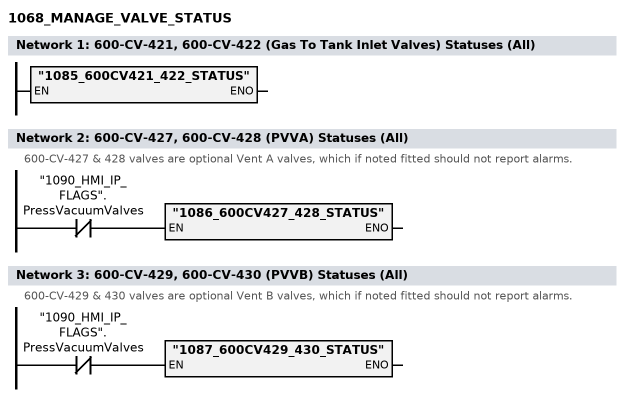
   RUNG wire#powerrail
      "1085_600CV421_422_STATUS"()
   END_RUNG
   // the same network as SCL:
   "1085_600CV421_422_STATUS"();
END_REGION

REGION Network 2: 600-CV-427, 600-CV-428 (PVVA) Statuses (All)
   // 600-CV-427 & 428 valves are optional Vent A valves, which if noted fitted should not report alarms.
   RUNG wire#powerrail
      I_Contact( "1090_HMI_IP_FLAGS".PressVacuumValves )
      "1086_600CV427_428_STATUS"()
   END_RUNG
   // the same network as SCL:
   IF NOT "1090_HMI_IP_FLAGS".PressVacuumValves THEN "1086_600CV427_428_STATUS"(); END_IF;
END_REGION

REGION Network 3: 600-CV-429, 600-CV-430 (PVVB) Statuses (All)
   // 600-CV-429 & 430 valves are optional Vent B valves, which if noted fitted should not report alarms.
   RUNG wire#powerrail
      I_Contact( "1090_HMI_IP_FLAGS".PressVacuumValves )
      "1087_600CV429_430_STATUS"()
   END_RUNG
   // the same network as SCL:
   IF NOT "1090_HMI_IP_FLAGS".PressVacuumValves THEN "1087_600CV429_430_STATUS"(); END_IF;
END_REGION
END_FUNCTION

// folder: 1000 - 1999 BWT System Control/1060 - 1089 Alarm & Valve Status Handling/1070 - 1079 Tank Alarms

FUNCTION "1070_LT421_422_ALARMS" : Void   // FC1070, LAD
{ S7_Optimized_Access := 'TRUE' }
VERSION : 0.1
// Alarm wrapper function for BWT Level on each tank.
// DummyIn and DummyAlarm are used to manage the unused I/O in the analog health trips function as this function only uses Low and High warnings, it does not output HighHigh or LowLow alarms.
   VAR_TEMP
      DummyIn : Real;   // Dummy input used if alarms are Low and High only.
      DummyAlarm : Bool;   // Dummy output used if alarms are Low and High only.
   END_VAR
BEGIN

REGION Network 1: LT421, LT422 Alarms (RIO 01: FPT. 1P, 1S)
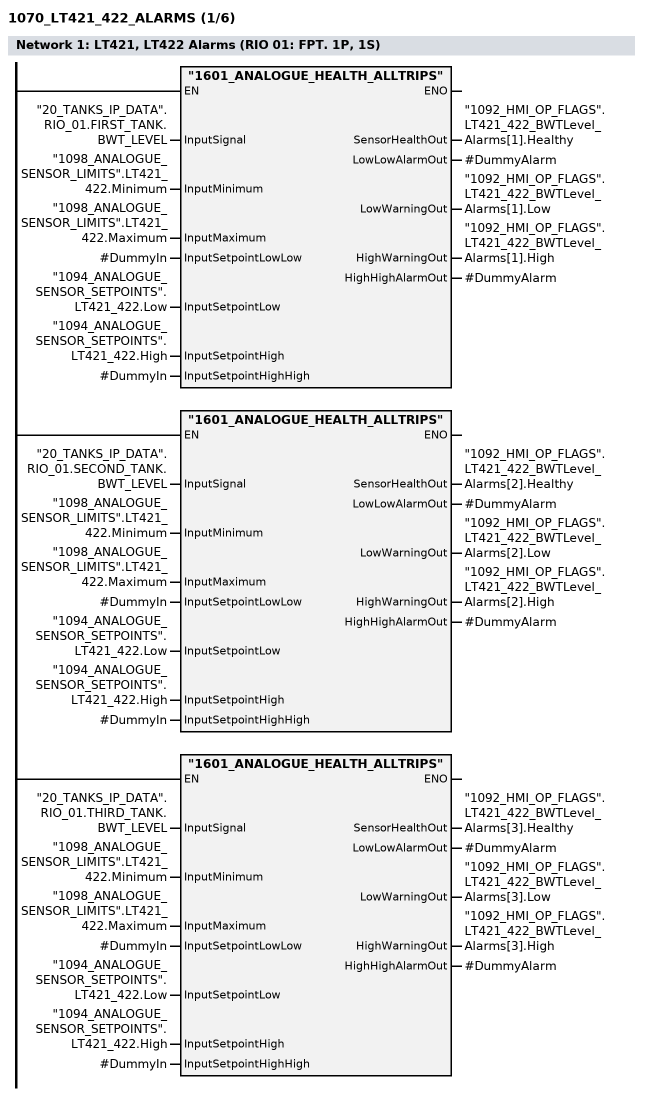
   RUNG wire#powerrail
      "1601_ANALOGUE_HEALTH_ALLTRIPS"(InputSignal := "20_TANKS_IP_DATA".RIO_01.FIRST_TANK.BWT_LEVEL, InputMinimum := "1098_ANALOGUE_SENSOR_LIMITS".LT421_422.Minimum, InputMaximum := "1098_ANALOGUE_SENSOR_LIMITS".LT421_422.Maximum, InputSetpointLowLow := #DummyIn, InputSetpointLow := "1094_ANALOGUE_SENSOR_SETPOINTS".LT421_422.Low, InputSetpointHigh := "1094_ANALOGUE_SENSOR_SETPOINTS".LT421_422.High, InputSetpointHighHigh := #DummyIn, SensorHealthOut => "1092_HMI_OP_FLAGS".LT421_422_BWTLevel_Alarms[1].Healthy, LowLowAlarmOut => #DummyAlarm, LowWarningOut => "1092_HMI_OP_FLAGS".LT421_422_BWTLevel_Alarms[1].Low, HighWarningOut => "1092_HMI_OP_FLAGS".LT421_422_BWTLevel_Alarms[1].High, HighHighAlarmOut => #DummyAlarm)
   END_RUNG
   RUNG wire#powerrail
      "1601_ANALOGUE_HEALTH_ALLTRIPS"(InputSignal := "20_TANKS_IP_DATA".RIO_01.SECOND_TANK.BWT_LEVEL, InputMinimum := "1098_ANALOGUE_SENSOR_LIMITS".LT421_422.Minimum, InputMaximum := "1098_ANALOGUE_SENSOR_LIMITS".LT421_422.Maximum, InputSetpointLowLow := #DummyIn, InputSetpointLow := "1094_ANALOGUE_SENSOR_SETPOINTS".LT421_422.Low, InputSetpointHigh := "1094_ANALOGUE_SENSOR_SETPOINTS".LT421_422.High, InputSetpointHighHigh := #DummyIn, SensorHealthOut => "1092_HMI_OP_FLAGS".LT421_422_BWTLevel_Alarms[2].Healthy, LowLowAlarmOut => #DummyAlarm, LowWarningOut => "1092_HMI_OP_FLAGS".LT421_422_BWTLevel_Alarms[2].Low, HighWarningOut => "1092_HMI_OP_FLAGS".LT421_422_BWTLevel_Alarms[2].High, HighHighAlarmOut => #DummyAlarm)
   END_RUNG
   RUNG wire#powerrail
      "1601_ANALOGUE_HEALTH_ALLTRIPS"(InputSignal := "20_TANKS_IP_DATA".RIO_01.THIRD_TANK.BWT_LEVEL, InputMinimum := "1098_ANALOGUE_SENSOR_LIMITS".LT421_422.Minimum, InputMaximum := "1098_ANALOGUE_SENSOR_LIMITS".LT421_422.Maximum, InputSetpointLowLow := #DummyIn, InputSetpointLow := "1094_ANALOGUE_SENSOR_SETPOINTS".LT421_422.Low, InputSetpointHigh := "1094_ANALOGUE_SENSOR_SETPOINTS".LT421_422.High, InputSetpointHighHigh := #DummyIn, SensorHealthOut => "1092_HMI_OP_FLAGS".LT421_422_BWTLevel_Alarms[3].Healthy, LowLowAlarmOut => #DummyAlarm, LowWarningOut => "1092_HMI_OP_FLAGS".LT421_422_BWTLevel_Alarms[3].Low, HighWarningOut => "1092_HMI_OP_FLAGS".LT421_422_BWTLevel_Alarms[3].High, HighHighAlarmOut => #DummyAlarm)
   END_RUNG
   // the same network as SCL:
   "1601_ANALOGUE_HEALTH_ALLTRIPS"(InputSignal := "20_TANKS_IP_DATA".RIO_01.FIRST_TANK.BWT_LEVEL,
                           InputMinimum := "1098_ANALOGUE_SENSOR_LIMITS".LT421_422.Minimum,
                           InputMaximum := "1098_ANALOGUE_SENSOR_LIMITS".LT421_422.Maximum,
                           InputSetpointLowLow := #DummyIn,
                           InputSetpointLow := "1094_ANALOGUE_SENSOR_SETPOINTS".LT421_422.Low,
                           InputSetpointHigh := "1094_ANALOGUE_SENSOR_SETPOINTS".LT421_422.High,
                           InputSetpointHighHigh := #DummyIn,
                           SensorHealthOut => "1092_HMI_OP_FLAGS".LT421_422_BWTLevel_Alarms[1].Healthy,
                           LowLowAlarmOut => #DummyAlarm,
                           LowWarningOut => "1092_HMI_OP_FLAGS".LT421_422_BWTLevel_Alarms[1].Low,
                           HighWarningOut => "1092_HMI_OP_FLAGS".LT421_422_BWTLevel_Alarms[1].High,
                           HighHighAlarmOut => #DummyAlarm);
   "1601_ANALOGUE_HEALTH_ALLTRIPS"(InputSignal := "20_TANKS_IP_DATA".RIO_01.SECOND_TANK.BWT_LEVEL,
                           InputMinimum := "1098_ANALOGUE_SENSOR_LIMITS".LT421_422.Minimum,
                           InputMaximum := "1098_ANALOGUE_SENSOR_LIMITS".LT421_422.Maximum,
                           InputSetpointLowLow := #DummyIn,
                           InputSetpointLow := "1094_ANALOGUE_SENSOR_SETPOINTS".LT421_422.Low,
                           InputSetpointHigh := "1094_ANALOGUE_SENSOR_SETPOINTS".LT421_422.High,
                           InputSetpointHighHigh := #DummyIn,
                           SensorHealthOut => "1092_HMI_OP_FLAGS".LT421_422_BWTLevel_Alarms[2].Healthy,
                           LowLowAlarmOut => #DummyAlarm,
                           LowWarningOut => "1092_HMI_OP_FLAGS".LT421_422_BWTLevel_Alarms[2].Low,
                           HighWarningOut => "1092_HMI_OP_FLAGS".LT421_422_BWTLevel_Alarms[2].High,
                           HighHighAlarmOut => #DummyAlarm);
   "1601_ANALOGUE_HEALTH_ALLTRIPS"(InputSignal := "20_TANKS_IP_DATA".RIO_01.THIRD_TANK.BWT_LEVEL,
                           InputMinimum := "1098_ANALOGUE_SENSOR_LIMITS".LT421_422.Minimum,
                           InputMaximum := "1098_ANALOGUE_SENSOR_LIMITS".LT421_422.Maximum,
                           InputSetpointLowLow := #DummyIn,
                           InputSetpointLow := "1094_ANALOGUE_SENSOR_SETPOINTS".LT421_422.Low,
                           InputSetpointHigh := "1094_ANALOGUE_SENSOR_SETPOINTS".LT421_422.High,
                           InputSetpointHighHigh := #DummyIn,
                           SensorHealthOut => "1092_HMI_OP_FLAGS".LT421_422_BWTLevel_Alarms[3].Healthy,
                           LowLowAlarmOut => #DummyAlarm,
                           LowWarningOut => "1092_HMI_OP_FLAGS".LT421_422_BWTLevel_Alarms[3].Low,
                           HighWarningOut => "1092_HMI_OP_FLAGS".LT421_422_BWTLevel_Alarms[3].High,
                           HighHighAlarmOut => #DummyAlarm);
END_REGION

REGION Network 2: LT421, LT422 Alarms (RIO 02: 2P, 2S)
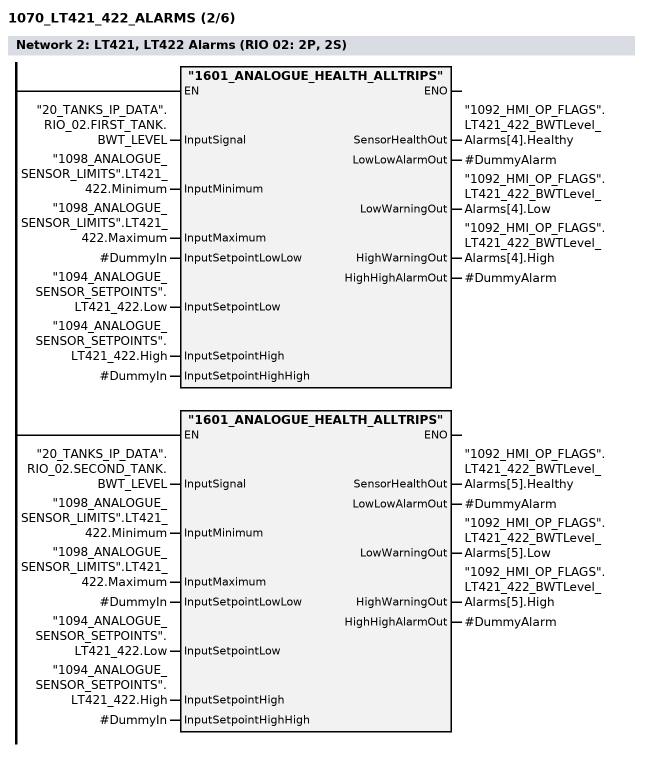
   RUNG wire#powerrail
      "1601_ANALOGUE_HEALTH_ALLTRIPS"(InputSignal := "20_TANKS_IP_DATA".RIO_02.FIRST_TANK.BWT_LEVEL, InputMinimum := "1098_ANALOGUE_SENSOR_LIMITS".LT421_422.Minimum, InputMaximum := "1098_ANALOGUE_SENSOR_LIMITS".LT421_422.Maximum, InputSetpointLowLow := #DummyIn, InputSetpointLow := "1094_ANALOGUE_SENSOR_SETPOINTS".LT421_422.Low, InputSetpointHigh := "1094_ANALOGUE_SENSOR_SETPOINTS".LT421_422.High, InputSetpointHighHigh := #DummyIn, SensorHealthOut => "1092_HMI_OP_FLAGS".LT421_422_BWTLevel_Alarms[4].Healthy, LowLowAlarmOut => #DummyAlarm, LowWarningOut => "1092_HMI_OP_FLAGS".LT421_422_BWTLevel_Alarms[4].Low, HighWarningOut => "1092_HMI_OP_FLAGS".LT421_422_BWTLevel_Alarms[4].High, HighHighAlarmOut => #DummyAlarm)
   END_RUNG
   RUNG wire#powerrail
      "1601_ANALOGUE_HEALTH_ALLTRIPS"(InputSignal := "20_TANKS_IP_DATA".RIO_02.SECOND_TANK.BWT_LEVEL, InputMinimum := "1098_ANALOGUE_SENSOR_LIMITS".LT421_422.Minimum, InputMaximum := "1098_ANALOGUE_SENSOR_LIMITS".LT421_422.Maximum, InputSetpointLowLow := #DummyIn, InputSetpointLow := "1094_ANALOGUE_SENSOR_SETPOINTS".LT421_422.Low, InputSetpointHigh := "1094_ANALOGUE_SENSOR_SETPOINTS".LT421_422.High, InputSetpointHighHigh := #DummyIn, SensorHealthOut => "1092_HMI_OP_FLAGS".LT421_422_BWTLevel_Alarms[5].Healthy, LowLowAlarmOut => #DummyAlarm, LowWarningOut => "1092_HMI_OP_FLAGS".LT421_422_BWTLevel_Alarms[5].Low, HighWarningOut => "1092_HMI_OP_FLAGS".LT421_422_BWTLevel_Alarms[5].High, HighHighAlarmOut => #DummyAlarm)
   END_RUNG
   // the same network as SCL:
   "1601_ANALOGUE_HEALTH_ALLTRIPS"(InputSignal := "20_TANKS_IP_DATA".RIO_02.FIRST_TANK.BWT_LEVEL,
                           InputMinimum := "1098_ANALOGUE_SENSOR_LIMITS".LT421_422.Minimum,
                           InputMaximum := "1098_ANALOGUE_SENSOR_LIMITS".LT421_422.Maximum,
                           InputSetpointLowLow := #DummyIn,
                           InputSetpointLow := "1094_ANALOGUE_SENSOR_SETPOINTS".LT421_422.Low,
                           InputSetpointHigh := "1094_ANALOGUE_SENSOR_SETPOINTS".LT421_422.High,
                           InputSetpointHighHigh := #DummyIn,
                           SensorHealthOut => "1092_HMI_OP_FLAGS".LT421_422_BWTLevel_Alarms[4].Healthy,
                           LowLowAlarmOut => #DummyAlarm,
                           LowWarningOut => "1092_HMI_OP_FLAGS".LT421_422_BWTLevel_Alarms[4].Low,
                           HighWarningOut => "1092_HMI_OP_FLAGS".LT421_422_BWTLevel_Alarms[4].High,
                           HighHighAlarmOut => #DummyAlarm);
   "1601_ANALOGUE_HEALTH_ALLTRIPS"(InputSignal := "20_TANKS_IP_DATA".RIO_02.SECOND_TANK.BWT_LEVEL,
                           InputMinimum := "1098_ANALOGUE_SENSOR_LIMITS".LT421_422.Minimum,
                           InputMaximum := "1098_ANALOGUE_SENSOR_LIMITS".LT421_422.Maximum,
                           InputSetpointLowLow := #DummyIn,
                           InputSetpointLow := "1094_ANALOGUE_SENSOR_SETPOINTS".LT421_422.Low,
                           InputSetpointHigh := "1094_ANALOGUE_SENSOR_SETPOINTS".LT421_422.High,
                           InputSetpointHighHigh := #DummyIn,
                           SensorHealthOut => "1092_HMI_OP_FLAGS".LT421_422_BWTLevel_Alarms[5].Healthy,
                           LowLowAlarmOut => #DummyAlarm,
                           LowWarningOut => "1092_HMI_OP_FLAGS".LT421_422_BWTLevel_Alarms[5].Low,
                           HighWarningOut => "1092_HMI_OP_FLAGS".LT421_422_BWTLevel_Alarms[5].High,
                           HighHighAlarmOut => #DummyAlarm);
END_REGION

REGION Network 3: LT421, LT422 Alarms (RIO 03: 3P, 3S)
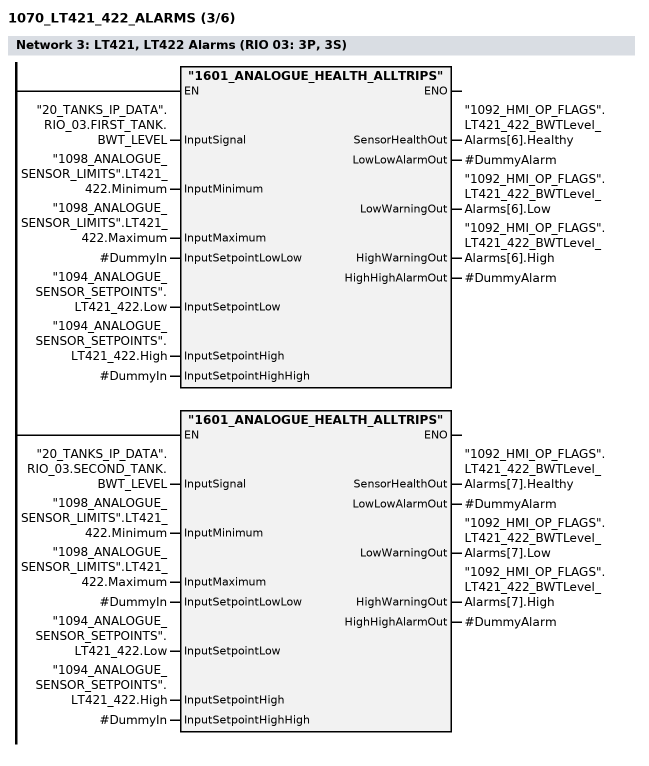
   RUNG wire#powerrail
      "1601_ANALOGUE_HEALTH_ALLTRIPS"(InputSignal := "20_TANKS_IP_DATA".RIO_03.FIRST_TANK.BWT_LEVEL, InputMinimum := "1098_ANALOGUE_SENSOR_LIMITS".LT421_422.Minimum, InputMaximum := "1098_ANALOGUE_SENSOR_LIMITS".LT421_422.Maximum, InputSetpointLowLow := #DummyIn, InputSetpointLow := "1094_ANALOGUE_SENSOR_SETPOINTS".LT421_422.Low, InputSetpointHigh := "1094_ANALOGUE_SENSOR_SETPOINTS".LT421_422.High, InputSetpointHighHigh := #DummyIn, SensorHealthOut => "1092_HMI_OP_FLAGS".LT421_422_BWTLevel_Alarms[6].Healthy, LowLowAlarmOut => #DummyAlarm, LowWarningOut => "1092_HMI_OP_FLAGS".LT421_422_BWTLevel_Alarms[6].Low, HighWarningOut => "1092_HMI_OP_FLAGS".LT421_422_BWTLevel_Alarms[6].High, HighHighAlarmOut => #DummyAlarm)
   END_RUNG
   RUNG wire#powerrail
      "1601_ANALOGUE_HEALTH_ALLTRIPS"(InputSignal := "20_TANKS_IP_DATA".RIO_03.SECOND_TANK.BWT_LEVEL, InputMinimum := "1098_ANALOGUE_SENSOR_LIMITS".LT421_422.Minimum, InputMaximum := "1098_ANALOGUE_SENSOR_LIMITS".LT421_422.Maximum, InputSetpointLowLow := #DummyIn, InputSetpointLow := "1094_ANALOGUE_SENSOR_SETPOINTS".LT421_422.Low, InputSetpointHigh := "1094_ANALOGUE_SENSOR_SETPOINTS".LT421_422.High, InputSetpointHighHigh := #DummyIn, SensorHealthOut => "1092_HMI_OP_FLAGS".LT421_422_BWTLevel_Alarms[7].Healthy, LowLowAlarmOut => #DummyAlarm, LowWarningOut => "1092_HMI_OP_FLAGS".LT421_422_BWTLevel_Alarms[7].Low, HighWarningOut => "1092_HMI_OP_FLAGS".LT421_422_BWTLevel_Alarms[7].High, HighHighAlarmOut => #DummyAlarm)
   END_RUNG
   // the same network as SCL:
   "1601_ANALOGUE_HEALTH_ALLTRIPS"(InputSignal := "20_TANKS_IP_DATA".RIO_03.FIRST_TANK.BWT_LEVEL,
                           InputMinimum := "1098_ANALOGUE_SENSOR_LIMITS".LT421_422.Minimum,
                           InputMaximum := "1098_ANALOGUE_SENSOR_LIMITS".LT421_422.Maximum,
                           InputSetpointLowLow := #DummyIn,
                           InputSetpointLow := "1094_ANALOGUE_SENSOR_SETPOINTS".LT421_422.Low,
                           InputSetpointHigh := "1094_ANALOGUE_SENSOR_SETPOINTS".LT421_422.High,
                           InputSetpointHighHigh := #DummyIn,
                           SensorHealthOut => "1092_HMI_OP_FLAGS".LT421_422_BWTLevel_Alarms[6].Healthy,
                           LowLowAlarmOut => #DummyAlarm,
                           LowWarningOut => "1092_HMI_OP_FLAGS".LT421_422_BWTLevel_Alarms[6].Low,
                           HighWarningOut => "1092_HMI_OP_FLAGS".LT421_422_BWTLevel_Alarms[6].High,
                           HighHighAlarmOut => #DummyAlarm);
   "1601_ANALOGUE_HEALTH_ALLTRIPS"(InputSignal := "20_TANKS_IP_DATA".RIO_03.SECOND_TANK.BWT_LEVEL,
                           InputMinimum := "1098_ANALOGUE_SENSOR_LIMITS".LT421_422.Minimum,
                           InputMaximum := "1098_ANALOGUE_SENSOR_LIMITS".LT421_422.Maximum,
                           InputSetpointLowLow := #DummyIn,
                           InputSetpointLow := "1094_ANALOGUE_SENSOR_SETPOINTS".LT421_422.Low,
                           InputSetpointHigh := "1094_ANALOGUE_SENSOR_SETPOINTS".LT421_422.High,
                           InputSetpointHighHigh := #DummyIn,
                           SensorHealthOut => "1092_HMI_OP_FLAGS".LT421_422_BWTLevel_Alarms[7].Healthy,
                           LowLowAlarmOut => #DummyAlarm,
                           LowWarningOut => "1092_HMI_OP_FLAGS".LT421_422_BWTLevel_Alarms[7].Low,
                           HighWarningOut => "1092_HMI_OP_FLAGS".LT421_422_BWTLevel_Alarms[7].High,
                           HighHighAlarmOut => #DummyAlarm);
END_REGION

REGION Network 4: LT421, LT422 Alarms (RIO 04: 4P, 4S)
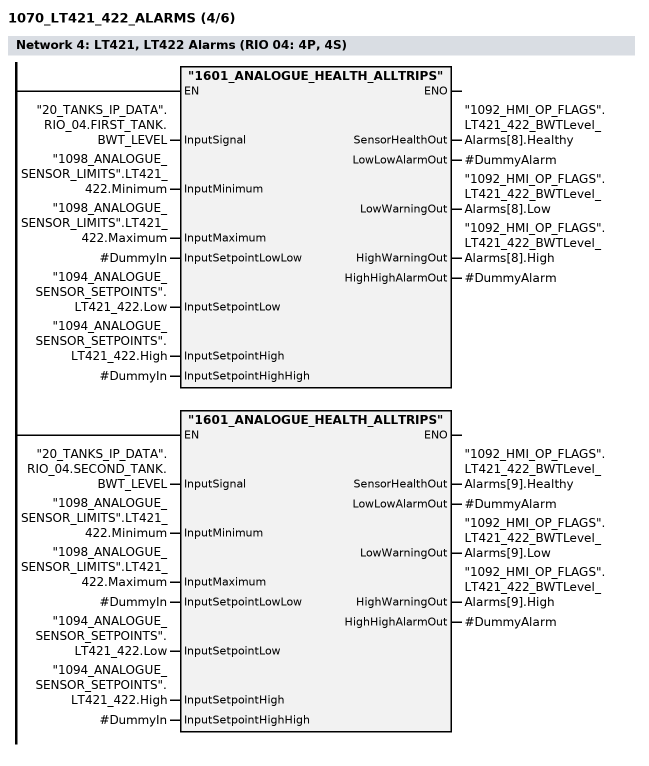
   RUNG wire#powerrail
      "1601_ANALOGUE_HEALTH_ALLTRIPS"(InputSignal := "20_TANKS_IP_DATA".RIO_04.FIRST_TANK.BWT_LEVEL, InputMinimum := "1098_ANALOGUE_SENSOR_LIMITS".LT421_422.Minimum, InputMaximum := "1098_ANALOGUE_SENSOR_LIMITS".LT421_422.Maximum, InputSetpointLowLow := #DummyIn, InputSetpointLow := "1094_ANALOGUE_SENSOR_SETPOINTS".LT421_422.Low, InputSetpointHigh := "1094_ANALOGUE_SENSOR_SETPOINTS".LT421_422.High, InputSetpointHighHigh := #DummyIn, SensorHealthOut => "1092_HMI_OP_FLAGS".LT421_422_BWTLevel_Alarms[8].Healthy, LowLowAlarmOut => #DummyAlarm, LowWarningOut => "1092_HMI_OP_FLAGS".LT421_422_BWTLevel_Alarms[8].Low, HighWarningOut => "1092_HMI_OP_FLAGS".LT421_422_BWTLevel_Alarms[8].High, HighHighAlarmOut => #DummyAlarm)
   END_RUNG
   RUNG wire#powerrail
      "1601_ANALOGUE_HEALTH_ALLTRIPS"(InputSignal := "20_TANKS_IP_DATA".RIO_04.SECOND_TANK.BWT_LEVEL, InputMinimum := "1098_ANALOGUE_SENSOR_LIMITS".LT421_422.Minimum, InputMaximum := "1098_ANALOGUE_SENSOR_LIMITS".LT421_422.Maximum, InputSetpointLowLow := #DummyIn, InputSetpointLow := "1094_ANALOGUE_SENSOR_SETPOINTS".LT421_422.Low, InputSetpointHigh := "1094_ANALOGUE_SENSOR_SETPOINTS".LT421_422.High, InputSetpointHighHigh := #DummyIn, SensorHealthOut => "1092_HMI_OP_FLAGS".LT421_422_BWTLevel_Alarms[9].Healthy, LowLowAlarmOut => #DummyAlarm, LowWarningOut => "1092_HMI_OP_FLAGS".LT421_422_BWTLevel_Alarms[9].Low, HighWarningOut => "1092_HMI_OP_FLAGS".LT421_422_BWTLevel_Alarms[9].High, HighHighAlarmOut => #DummyAlarm)
   END_RUNG
   // the same network as SCL:
   "1601_ANALOGUE_HEALTH_ALLTRIPS"(InputSignal := "20_TANKS_IP_DATA".RIO_04.FIRST_TANK.BWT_LEVEL,
                           InputMinimum := "1098_ANALOGUE_SENSOR_LIMITS".LT421_422.Minimum,
                           InputMaximum := "1098_ANALOGUE_SENSOR_LIMITS".LT421_422.Maximum,
                           InputSetpointLowLow := #DummyIn,
                           InputSetpointLow := "1094_ANALOGUE_SENSOR_SETPOINTS".LT421_422.Low,
                           InputSetpointHigh := "1094_ANALOGUE_SENSOR_SETPOINTS".LT421_422.High,
                           InputSetpointHighHigh := #DummyIn,
                           SensorHealthOut => "1092_HMI_OP_FLAGS".LT421_422_BWTLevel_Alarms[8].Healthy,
                           LowLowAlarmOut => #DummyAlarm,
                           LowWarningOut => "1092_HMI_OP_FLAGS".LT421_422_BWTLevel_Alarms[8].Low,
                           HighWarningOut => "1092_HMI_OP_FLAGS".LT421_422_BWTLevel_Alarms[8].High,
                           HighHighAlarmOut => #DummyAlarm);
   "1601_ANALOGUE_HEALTH_ALLTRIPS"(InputSignal := "20_TANKS_IP_DATA".RIO_04.SECOND_TANK.BWT_LEVEL,
                           InputMinimum := "1098_ANALOGUE_SENSOR_LIMITS".LT421_422.Minimum,
                           InputMaximum := "1098_ANALOGUE_SENSOR_LIMITS".LT421_422.Maximum,
                           InputSetpointLowLow := #DummyIn,
                           InputSetpointLow := "1094_ANALOGUE_SENSOR_SETPOINTS".LT421_422.Low,
                           InputSetpointHigh := "1094_ANALOGUE_SENSOR_SETPOINTS".LT421_422.High,
                           InputSetpointHighHigh := #DummyIn,
                           SensorHealthOut => "1092_HMI_OP_FLAGS".LT421_422_BWTLevel_Alarms[9].Healthy,
                           LowLowAlarmOut => #DummyAlarm,
                           LowWarningOut => "1092_HMI_OP_FLAGS".LT421_422_BWTLevel_Alarms[9].Low,
                           HighWarningOut => "1092_HMI_OP_FLAGS".LT421_422_BWTLevel_Alarms[9].High,
                           HighHighAlarmOut => #DummyAlarm);
END_REGION

REGION Network 5: LT421, LT422 Alarms (RIO 05: 5P, 5S)
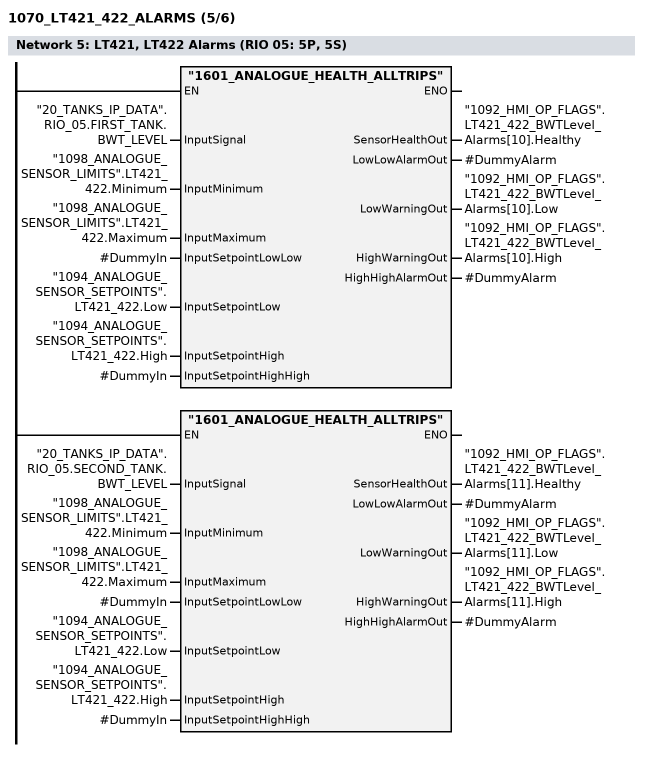
   RUNG wire#powerrail
      "1601_ANALOGUE_HEALTH_ALLTRIPS"(InputSignal := "20_TANKS_IP_DATA".RIO_05.FIRST_TANK.BWT_LEVEL, InputMinimum := "1098_ANALOGUE_SENSOR_LIMITS".LT421_422.Minimum, InputMaximum := "1098_ANALOGUE_SENSOR_LIMITS".LT421_422.Maximum, InputSetpointLowLow := #DummyIn, InputSetpointLow := "1094_ANALOGUE_SENSOR_SETPOINTS".LT421_422.Low, InputSetpointHigh := "1094_ANALOGUE_SENSOR_SETPOINTS".LT421_422.High, InputSetpointHighHigh := #DummyIn, SensorHealthOut => "1092_HMI_OP_FLAGS".LT421_422_BWTLevel_Alarms[10].Healthy, LowLowAlarmOut => #DummyAlarm, LowWarningOut => "1092_HMI_OP_FLAGS".LT421_422_BWTLevel_Alarms[10].Low, HighWarningOut => "1092_HMI_OP_FLAGS".LT421_422_BWTLevel_Alarms[10].High, HighHighAlarmOut => #DummyAlarm)
   END_RUNG
   RUNG wire#powerrail
      "1601_ANALOGUE_HEALTH_ALLTRIPS"(InputSignal := "20_TANKS_IP_DATA".RIO_05.SECOND_TANK.BWT_LEVEL, InputMinimum := "1098_ANALOGUE_SENSOR_LIMITS".LT421_422.Minimum, InputMaximum := "1098_ANALOGUE_SENSOR_LIMITS".LT421_422.Maximum, InputSetpointLowLow := #DummyIn, InputSetpointLow := "1094_ANALOGUE_SENSOR_SETPOINTS".LT421_422.Low, InputSetpointHigh := "1094_ANALOGUE_SENSOR_SETPOINTS".LT421_422.High, InputSetpointHighHigh := #DummyIn, SensorHealthOut => "1092_HMI_OP_FLAGS".LT421_422_BWTLevel_Alarms[11].Healthy, LowLowAlarmOut => #DummyAlarm, LowWarningOut => "1092_HMI_OP_FLAGS".LT421_422_BWTLevel_Alarms[11].Low, HighWarningOut => "1092_HMI_OP_FLAGS".LT421_422_BWTLevel_Alarms[11].High, HighHighAlarmOut => #DummyAlarm)
   END_RUNG
   // the same network as SCL:
   "1601_ANALOGUE_HEALTH_ALLTRIPS"(InputSignal := "20_TANKS_IP_DATA".RIO_05.FIRST_TANK.BWT_LEVEL,
                           InputMinimum := "1098_ANALOGUE_SENSOR_LIMITS".LT421_422.Minimum,
                           InputMaximum := "1098_ANALOGUE_SENSOR_LIMITS".LT421_422.Maximum,
                           InputSetpointLowLow := #DummyIn,
                           InputSetpointLow := "1094_ANALOGUE_SENSOR_SETPOINTS".LT421_422.Low,
                           InputSetpointHigh := "1094_ANALOGUE_SENSOR_SETPOINTS".LT421_422.High,
                           InputSetpointHighHigh := #DummyIn,
                           SensorHealthOut => "1092_HMI_OP_FLAGS".LT421_422_BWTLevel_Alarms[10].Healthy,
                           LowLowAlarmOut => #DummyAlarm,
                           LowWarningOut => "1092_HMI_OP_FLAGS".LT421_422_BWTLevel_Alarms[10].Low,
                           HighWarningOut => "1092_HMI_OP_FLAGS".LT421_422_BWTLevel_Alarms[10].High,
                           HighHighAlarmOut => #DummyAlarm);
   "1601_ANALOGUE_HEALTH_ALLTRIPS"(InputSignal := "20_TANKS_IP_DATA".RIO_05.SECOND_TANK.BWT_LEVEL,
                           InputMinimum := "1098_ANALOGUE_SENSOR_LIMITS".LT421_422.Minimum,
                           InputMaximum := "1098_ANALOGUE_SENSOR_LIMITS".LT421_422.Maximum,
                           InputSetpointLowLow := #DummyIn,
                           InputSetpointLow := "1094_ANALOGUE_SENSOR_SETPOINTS".LT421_422.Low,
                           InputSetpointHigh := "1094_ANALOGUE_SENSOR_SETPOINTS".LT421_422.High,
                           InputSetpointHighHigh := #DummyIn,
                           SensorHealthOut => "1092_HMI_OP_FLAGS".LT421_422_BWTLevel_Alarms[11].Healthy,
                           LowLowAlarmOut => #DummyAlarm,
                           LowWarningOut => "1092_HMI_OP_FLAGS".LT421_422_BWTLevel_Alarms[11].Low,
                           HighWarningOut => "1092_HMI_OP_FLAGS".LT421_422_BWTLevel_Alarms[11].High,
                           HighHighAlarmOut => #DummyAlarm);
END_REGION

REGION Network 6: LT421, LT422 Alarms (RIO 06: 6P, 6S)
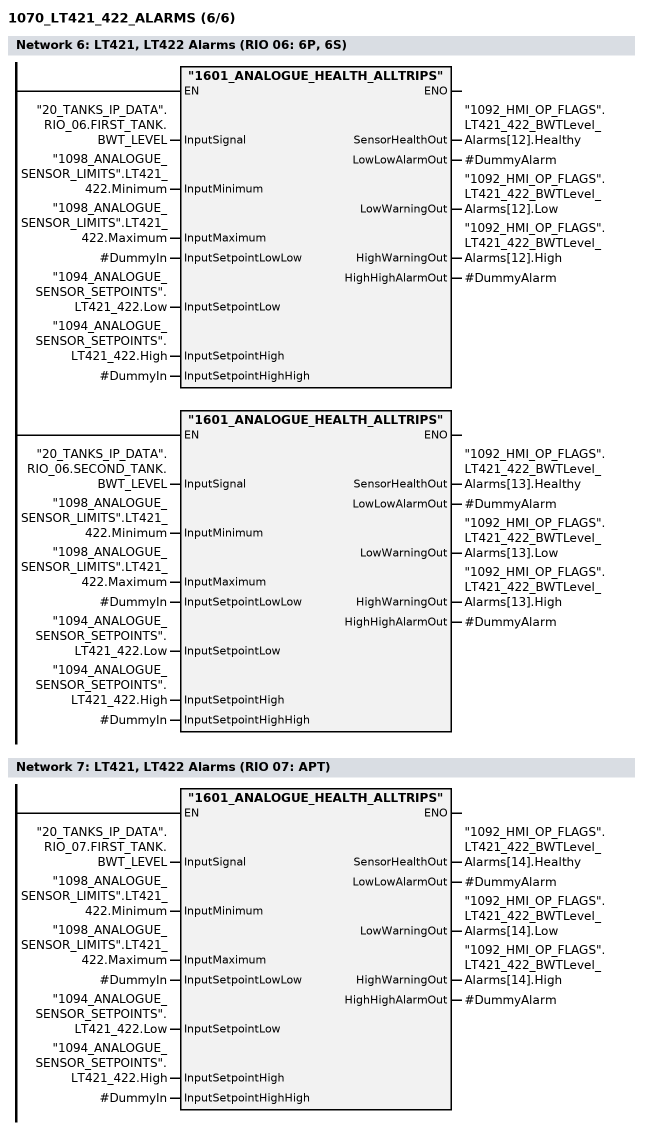
   RUNG wire#powerrail
      "1601_ANALOGUE_HEALTH_ALLTRIPS"(InputSignal := "20_TANKS_IP_DATA".RIO_06.FIRST_TANK.BWT_LEVEL, InputMinimum := "1098_ANALOGUE_SENSOR_LIMITS".LT421_422.Minimum, InputMaximum := "1098_ANALOGUE_SENSOR_LIMITS".LT421_422.Maximum, InputSetpointLowLow := #DummyIn, InputSetpointLow := "1094_ANALOGUE_SENSOR_SETPOINTS".LT421_422.Low, InputSetpointHigh := "1094_ANALOGUE_SENSOR_SETPOINTS".LT421_422.High, InputSetpointHighHigh := #DummyIn, SensorHealthOut => "1092_HMI_OP_FLAGS".LT421_422_BWTLevel_Alarms[12].Healthy, LowLowAlarmOut => #DummyAlarm, LowWarningOut => "1092_HMI_OP_FLAGS".LT421_422_BWTLevel_Alarms[12].Low, HighWarningOut => "1092_HMI_OP_FLAGS".LT421_422_BWTLevel_Alarms[12].High, HighHighAlarmOut => #DummyAlarm)
   END_RUNG
   RUNG wire#powerrail
      "1601_ANALOGUE_HEALTH_ALLTRIPS"(InputSignal := "20_TANKS_IP_DATA".RIO_06.SECOND_TANK.BWT_LEVEL, InputMinimum := "1098_ANALOGUE_SENSOR_LIMITS".LT421_422.Minimum, InputMaximum := "1098_ANALOGUE_SENSOR_LIMITS".LT421_422.Maximum, InputSetpointLowLow := #DummyIn, InputSetpointLow := "1094_ANALOGUE_SENSOR_SETPOINTS".LT421_422.Low, InputSetpointHigh := "1094_ANALOGUE_SENSOR_SETPOINTS".LT421_422.High, InputSetpointHighHigh := #DummyIn, SensorHealthOut => "1092_HMI_OP_FLAGS".LT421_422_BWTLevel_Alarms[13].Healthy, LowLowAlarmOut => #DummyAlarm, LowWarningOut => "1092_HMI_OP_FLAGS".LT421_422_BWTLevel_Alarms[13].Low, HighWarningOut => "1092_HMI_OP_FLAGS".LT421_422_BWTLevel_Alarms[13].High, HighHighAlarmOut => #DummyAlarm)
   END_RUNG
   // the same network as SCL:
   "1601_ANALOGUE_HEALTH_ALLTRIPS"(InputSignal := "20_TANKS_IP_DATA".RIO_06.FIRST_TANK.BWT_LEVEL,
                           InputMinimum := "1098_ANALOGUE_SENSOR_LIMITS".LT421_422.Minimum,
                           InputMaximum := "1098_ANALOGUE_SENSOR_LIMITS".LT421_422.Maximum,
                           InputSetpointLowLow := #DummyIn,
                           InputSetpointLow := "1094_ANALOGUE_SENSOR_SETPOINTS".LT421_422.Low,
                           InputSetpointHigh := "1094_ANALOGUE_SENSOR_SETPOINTS".LT421_422.High,
                           InputSetpointHighHigh := #DummyIn,
                           SensorHealthOut => "1092_HMI_OP_FLAGS".LT421_422_BWTLevel_Alarms[12].Healthy,
                           LowLowAlarmOut => #DummyAlarm,
                           LowWarningOut => "1092_HMI_OP_FLAGS".LT421_422_BWTLevel_Alarms[12].Low,
                           HighWarningOut => "1092_HMI_OP_FLAGS".LT421_422_BWTLevel_Alarms[12].High,
                           HighHighAlarmOut => #DummyAlarm);
   "1601_ANALOGUE_HEALTH_ALLTRIPS"(InputSignal := "20_TANKS_IP_DATA".RIO_06.SECOND_TANK.BWT_LEVEL,
                           InputMinimum := "1098_ANALOGUE_SENSOR_LIMITS".LT421_422.Minimum,
                           InputMaximum := "1098_ANALOGUE_SENSOR_LIMITS".LT421_422.Maximum,
                           InputSetpointLowLow := #DummyIn,
                           InputSetpointLow := "1094_ANALOGUE_SENSOR_SETPOINTS".LT421_422.Low,
                           InputSetpointHigh := "1094_ANALOGUE_SENSOR_SETPOINTS".LT421_422.High,
                           InputSetpointHighHigh := #DummyIn,
                           SensorHealthOut => "1092_HMI_OP_FLAGS".LT421_422_BWTLevel_Alarms[13].Healthy,
                           LowLowAlarmOut => #DummyAlarm,
                           LowWarningOut => "1092_HMI_OP_FLAGS".LT421_422_BWTLevel_Alarms[13].Low,
                           HighWarningOut => "1092_HMI_OP_FLAGS".LT421_422_BWTLevel_Alarms[13].High,
                           HighHighAlarmOut => #DummyAlarm);
END_REGION

REGION Network 7: LT421, LT422 Alarms (RIO 07: APT)
   RUNG wire#powerrail
      "1601_ANALOGUE_HEALTH_ALLTRIPS"(InputSignal := "20_TANKS_IP_DATA".RIO_07.FIRST_TANK.BWT_LEVEL, InputMinimum := "1098_ANALOGUE_SENSOR_LIMITS".LT421_422.Minimum, InputMaximum := "1098_ANALOGUE_SENSOR_LIMITS".LT421_422.Maximum, InputSetpointLowLow := #DummyIn, InputSetpointLow := "1094_ANALOGUE_SENSOR_SETPOINTS".LT421_422.Low, InputSetpointHigh := "1094_ANALOGUE_SENSOR_SETPOINTS".LT421_422.High, InputSetpointHighHigh := #DummyIn, SensorHealthOut => "1092_HMI_OP_FLAGS".LT421_422_BWTLevel_Alarms[14].Healthy, LowLowAlarmOut => #DummyAlarm, LowWarningOut => "1092_HMI_OP_FLAGS".LT421_422_BWTLevel_Alarms[14].Low, HighWarningOut => "1092_HMI_OP_FLAGS".LT421_422_BWTLevel_Alarms[14].High, HighHighAlarmOut => #DummyAlarm)
   END_RUNG
   // the same network as SCL:
   "1601_ANALOGUE_HEALTH_ALLTRIPS"(InputSignal := "20_TANKS_IP_DATA".RIO_07.FIRST_TANK.BWT_LEVEL,
                           InputMinimum := "1098_ANALOGUE_SENSOR_LIMITS".LT421_422.Minimum,
                           InputMaximum := "1098_ANALOGUE_SENSOR_LIMITS".LT421_422.Maximum,
                           InputSetpointLowLow := #DummyIn,
                           InputSetpointLow := "1094_ANALOGUE_SENSOR_SETPOINTS".LT421_422.Low,
                           InputSetpointHigh := "1094_ANALOGUE_SENSOR_SETPOINTS".LT421_422.High,
                           InputSetpointHighHigh := #DummyIn,
                           SensorHealthOut => "1092_HMI_OP_FLAGS".LT421_422_BWTLevel_Alarms[14].Healthy,
                           LowLowAlarmOut => #DummyAlarm,
                           LowWarningOut => "1092_HMI_OP_FLAGS".LT421_422_BWTLevel_Alarms[14].Low,
                           HighWarningOut => "1092_HMI_OP_FLAGS".LT421_422_BWTLevel_Alarms[14].High,
                           HighHighAlarmOut => #DummyAlarm);
END_REGION
END_FUNCTION

FUNCTION "1071_FIT417_418_ALARMS" : Void   // FC1071, LAD
{ S7_Optimized_Access := 'TRUE' }
VERSION : 0.1
// Alarm wrapper function for USD Flow on each tank.
BEGIN

REGION Network 1: FIT417, FIT418 Alarms (RIO 01: FPT. 1P, 1S)